// TIA Portal project "EdgeHowTos" (V16) (continued)
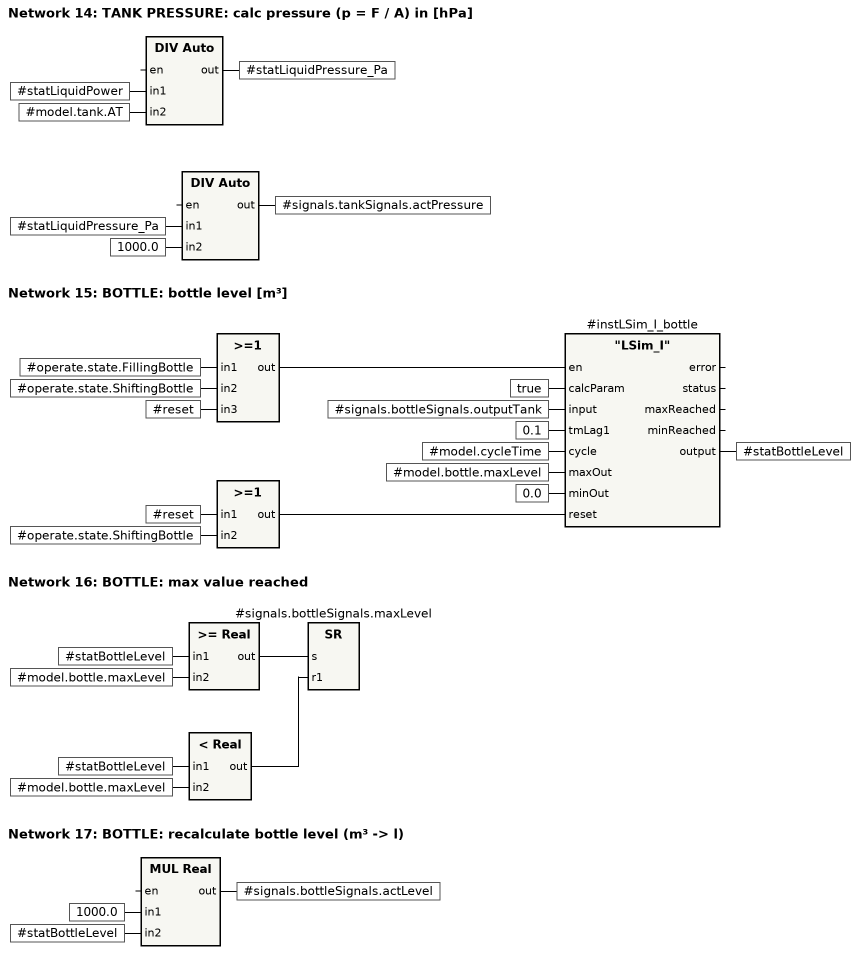
   #statLiquidPressure_Pa := #statLiquidPower / #model.tank.AT;
   #signals.tankSignals.actPressure := #statLiquidPressure_Pa / 1000.0;
END_REGION

REGION Network 15: BOTTLE: bottle level [m³]
   IF #operate.state.FillingBottle OR #operate.state.ShiftingBottle OR #reset THEN
       #instLSim_I_bottle(calcParam := true,   // "LSim_I"
                          input := #signals.bottleSignals.outputTank,
                          tmLag1 := 0.1,
                          cycle := #model.cycleTime,
                          maxOut := #model.bottle.maxLevel,
                          minOut := 0.0,
                          reset := #reset OR #operate.state.ShiftingBottle,
                          output => #statBottleLevel);
   END_IF;
END_REGION

REGION Network 16: BOTTLE: max value reached
   IF #statBottleLevel >= #model.bottle.maxLevel THEN
       #signals.bottleSignals.maxLevel := TRUE;   // SR flip-flop
   END_IF;
   IF #statBottleLevel < #model.bottle.maxLevel THEN #signals.bottleSignals.maxLevel := FALSE; END_IF;
END_REGION

REGION Network 17: BOTTLE: recalculate bottle level (m³ -> l)
   #signals.bottleSignals.actLevel := 1000.0 * #statBottleLevel;
END_REGION

REGION Network 18: HEAT: set init values
   // default value (statHeatingActive = false)
   // - temp = 20°C
   // - tmLag = 0.01
   // (set PT1 controller to initial temperature, otherwise PT1 controller would always start at 0°C)
   // 
   // heating phase (statHeatingActive = true)
   // - temp = 80°C
   // - tmLag = 1
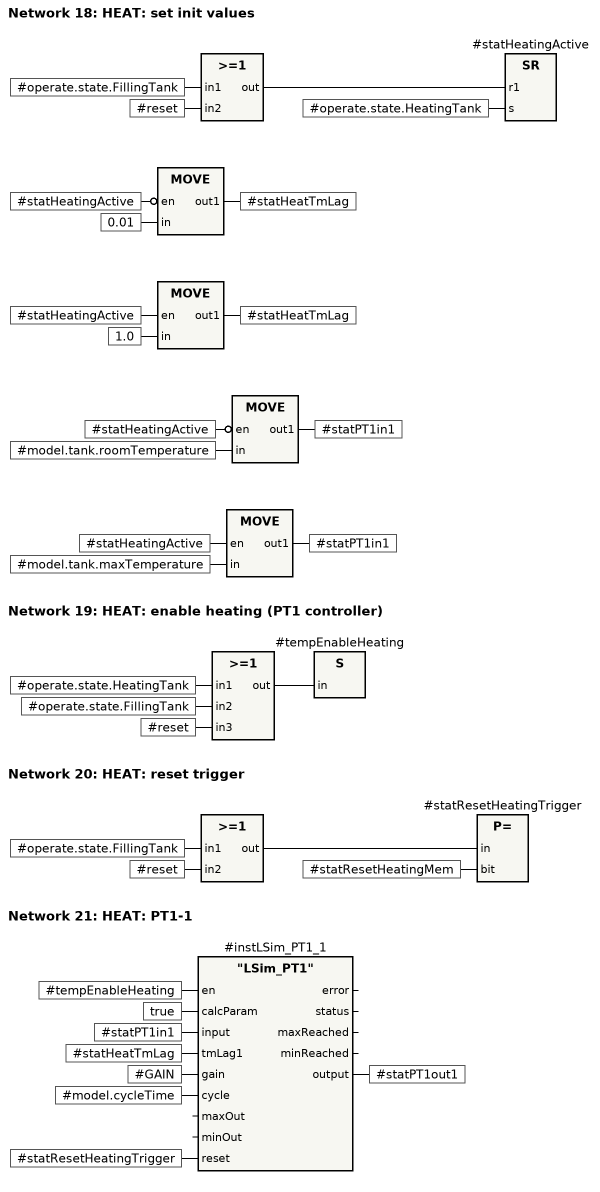
   IF #operate.state.HeatingTank THEN
       #statHeatingActive := TRUE;   // SR flip-flop
   END_IF;
   IF #operate.state.FillingTank OR #reset THEN #statHeatingActive := FALSE; END_IF;
   IF NOT #statHeatingActive THEN #statHeatTmLag := 0.01; END_IF;
   IF #statHeatingActive THEN #statHeatTmLag := 1.0; END_IF;
   IF NOT #statHeatingActive THEN #statPT1in1 := #model.tank.roomTemperature; END_IF;
   IF #statHeatingActive THEN #statPT1in1 := #model.tank.maxTemperature; END_IF;
END_REGION

REGION Network 19: HEAT: enable heating (PT1 controller)
   IF #operate.state.HeatingTank OR #operate.state.FillingTank OR #reset THEN
       #tempEnableHeating := TRUE;
   END_IF;
END_REGION

REGION Network 20: HEAT: reset trigger
   #_w1 := #operate.state.FillingTank OR #reset;
   #statResetHeatingTrigger := #_w1 AND NOT #statResetHeatingMem;   // rising edge
   #statResetHeatingMem := #_w1;
END_REGION

REGION Network 21: HEAT: PT1-1
   IF #tempEnableHeating THEN
       #instLSim_PT1_1(calcParam := true,   // "LSim_PT1"
                       input := #statPT1in1,
                       tmLag1 := #statHeatTmLag,
                       gain := #GAIN,
                       cycle := #model.cycleTime,
                       reset := #statResetHeatingTrigger,
                       output => #statPT1out1);
   END_IF;
END_REGION

REGION Network 22: HEAT: PT1-2
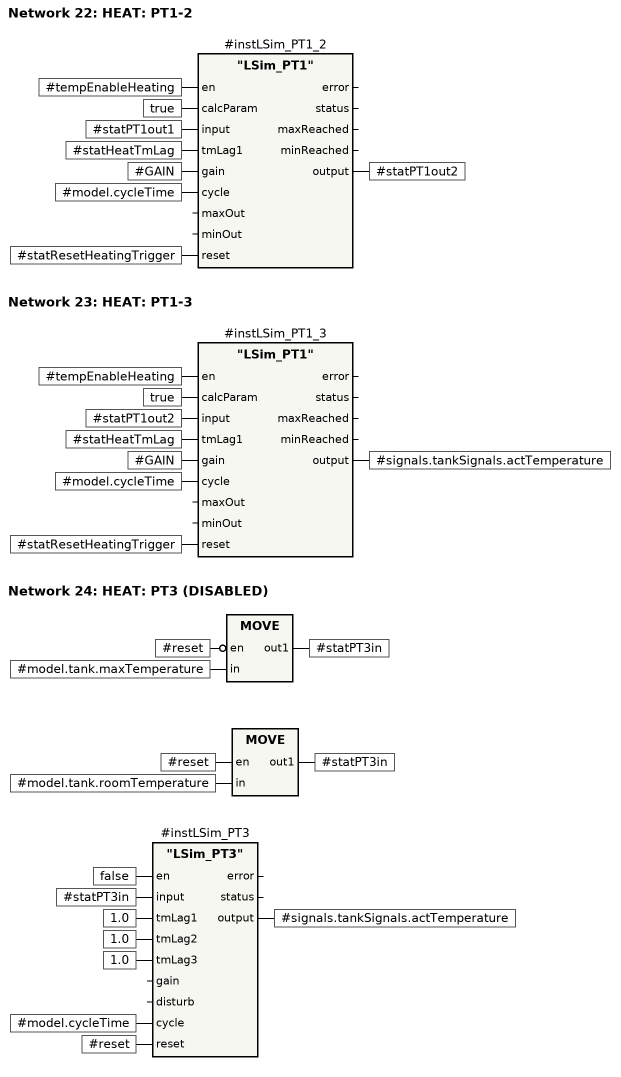
   IF #tempEnableHeating THEN
       #instLSim_PT1_2(calcParam := true,   // "LSim_PT1"
                       input := #statPT1out1,
                       tmLag1 := #statHeatTmLag,
                       gain := #GAIN,
                       cycle := #model.cycleTime,
                       reset := #statResetHeatingTrigger,
                       output => #statPT1out2);
   END_IF;
END_REGION

REGION Network 23: HEAT: PT1-3
   IF #tempEnableHeating THEN
       #instLSim_PT1_3(calcParam := true,   // "LSim_PT1"
                       input := #statPT1out2,
                       tmLag1 := #statHeatTmLag,
                       gain := #GAIN,
                       cycle := #model.cycleTime,
                       reset := #statResetHeatingTrigger,
                       output => #signals.tankSignals.actTemperature);
   END_IF;
END_REGION

REGION Network 24: HEAT: PT3 (DISABLED)
   IF NOT #reset THEN #statPT3in := #model.tank.maxTemperature; END_IF;
   IF #reset THEN #statPT3in := #model.tank.roomTemperature; END_IF;
   IF false THEN
       #instLSim_PT3(input := #statPT3in,   // "LSim_PT3"
                     tmLag1 := 1.0,
                     tmLag2 := 1.0,
                     tmLag3 := 1.0,
                     cycle := #model.cycleTime,
                     reset := #reset,
                     output => #signals.tankSignals.actTemperature);
   END_IF;
END_REGION

REGION Network 25: HEAT: max value reached
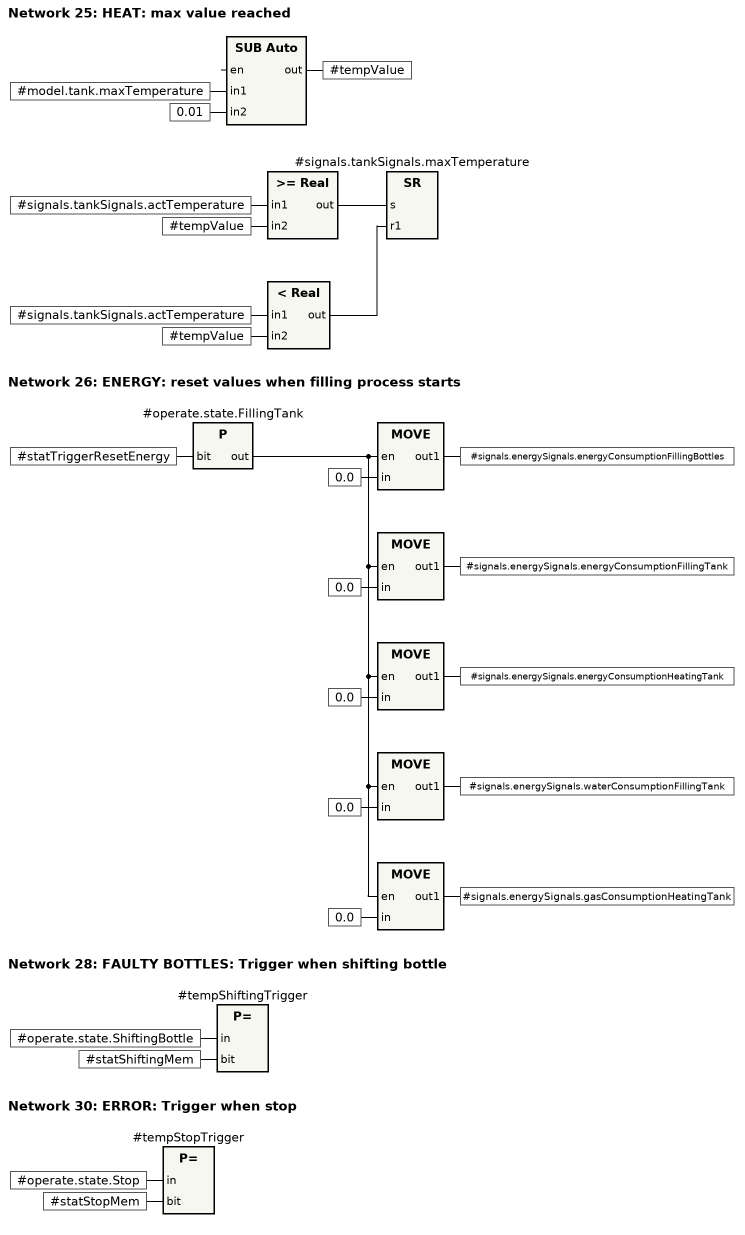
   #tempValue := #model.tank.maxTemperature - 0.01;
   IF #signals.tankSignals.actTemperature >= #tempValue THEN
       #signals.tankSignals.maxTemperature := TRUE;   // SR flip-flop
   END_IF;
   IF #signals.tankSignals.actTemperature < #tempValue THEN
       #signals.tankSignals.maxTemperature := FALSE;
   END_IF;
END_REGION

REGION Network 26: ENERGY: reset values when filling process starts
   #_w1 := #operate.state.FillingTank AND NOT #statTriggerResetEnergy;   // rising edge of #operate.state.FillingTank
   #statTriggerResetEnergy := #operate.state.FillingTank;
   IF #_w1 THEN
       #signals.energySignals.energyConsumptionFillingBottles := 0.0;
       #signals.energySignals.energyConsumptionFillingTank := 0.0;
       #signals.energySignals.energyConsumptionHeatingTank := 0.0;
       #signals.energySignals.waterConsumptionFillingTank := 0.0;
       #signals.energySignals.gasConsumptionHeatingTank := 0.0;
   END_IF;
END_REGION

REGION Network 27 (SCL): ENERGY: calculate values
   // generate random values for energy / water / gas consumption
   // energy [Wh] and water [l] consumption during filling tank
   // ----------------------------------------------------------
   IF #operate.state.FillingTank THEN
       "Random_Number"(Min := 10,
                       Max := 20,
                       RandomNumber => #tempRandomNumber);
       #tempRandomNumber := #tempRandomNumber / 100;
       #signals.energySignals.energyConsumptionFillingTank := #signals.energySignals.energyConsumptionFillingTank + #tempRandomNumber;
       #signals.energySignals.waterConsumptionFillingTank := #signals.tankSignals.actLevel;
   END_IF;

   // energy and gas consumption during heating tank [Wh]
   // ---------------------------------------------------
   IF #operate.state.HeatingTank THEN
       "Random_Number"(Min := 1,
                       Max := 8,
                       RandomNumber => #tempRandomNumber1);
       #tempRandomNumber1 := #tempRandomNumber1 / 10;
       #signals.energySignals.energyConsumptionHeatingTank := #signals.energySignals.energyConsumptionHeatingTank + #tempRandomNumber1;
       #signals.energySignals.gasConsumptionHeatingTank := #signals.energySignals.gasConsumptionHeatingTank + (#tempRandomNumber1 * 1.5);
   END_IF;

   // energy consumption during filling bottles [Wh]
   // -----------------------------------------------
   IF #operate.state.FillingBottle OR #operate.state.ShiftingBottle THEN
       "Random_Number"(Min := 10,
                       Max := 50,
                       RandomNumber => #tempRandomNumber2);
       #tempRandomNumber2 := #tempRandomNumber2 / 100;
       #signals.energySignals.energyConsumptionFillingBottles := #signals.energySignals.energyConsumptionFillingBottles + #tempRandomNumber2;
   END_IF;
END_REGION

REGION Network 28: FAULTY BOTTLES: Trigger when shifting bottle
   #tempShiftingTrigger := #operate.state.ShiftingBottle AND NOT #statShiftingMem;   // rising edge
   #statShiftingMem := #operate.state.ShiftingBottle;
END_REGION

REGION Network 29 (SCL): FAULTY BOTTLES: Simulate faulty bottles (generate random number)
   IF #tempShiftingTrigger THEN
       "Random_Number"(Min := 0,
                       Max := 8,
                       RandomNumber => #tempRandomNumber3);

       IF (#tempRandomNumber3 = 1) OR (#tempRandomNumber3 = 5) THEN
           #process.numberFaulty := #process.numberFaulty + 1;
       END_IF;

   END_IF;
END_REGION

REGION Network 30: ERROR: Trigger when stop
   #tempStopTrigger := #operate.state.Stop AND NOT #statStopMem;   // rising edge
   #statStopMem := #operate.state.Stop;
END_REGION

REGION Network 31 (SCL): ERROR: Simulate error
       IF #errors.errorSimulation THEN

           // random error generation
           IF #tempShiftingTrigger THEN
               "Random_Number"(Min := 0,
                               Max := 100,
                               RandomNumber => #tempRandomNumber5);

               // go into error state
               IF #tempRandomNumber5 = 1 THEN
                   #appSignals.APP_Error := true;
               END_IF;

           END_IF;

           // triggered error genertion
           IF #errors.errorTrigger THEN
               #appSignals.APP_Error := true;
           END_IF;


           // if timer finished (negative edge on it's output), go in stop > start again
           "F_TRIG_DB_Error_Finished"(CLK := #instTimerError.Q,
                                      Q => #statResetError);

           // reset error > machine goes automatically into stop
           IF #statResetError THEN
               #appSignals.APP_Error := false;
               #errors.errorCode := "ERROR_0_NO";
               #statResetError := false;
               #statStart := true;
           END_IF;

           IF #tempStopTrigger AND #statStart THEN
               #appSignals.APP_Start := true;
               #statStart := false;
           END_IF;

       END_IF;
END_REGION

REGION Network 32: ERROR: Trigger when new error comes in and start timer
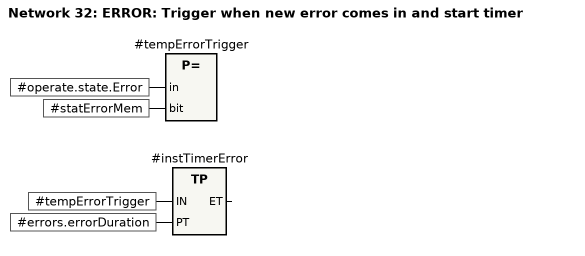
   #tempErrorTrigger := #operate.state.Error AND NOT #statErrorMem;   // rising edge
   #statErrorMem := #operate.state.Error;
   #instTimerError.TP(IN := #tempErrorTrigger, PT := #errors.errorDuration);
END_REGION

REGION Network 33 (SCL): ERROR: Simulate error codes
   // Codes btw. 1-6 (7 = HMI error)
   IF #errors.errorSimulation THEN

       // generate random error code
       IF #tempErrorTrigger AND (#errors.errorCode = "ERROR_0_NO") THEN

           "Random_Number"(Min := 1,
                           Max := 6,
                           RandomNumber => #tempRandomNumber4);

           #errors.errorCode := #tempRandomNumber4;

       END_IF;

   END_IF;
END_REGION
END_FUNCTION_BLOCK

FUNCTION_BLOCK "LSim_PT1"   // FB50, SCL
{ S7_Optimized_Access := 'TRUE' }
VERSION : 2.01
   VAR_INPUT
      calcParam : Bool;   // recalculate with new parameters
      input : Real;   // input signal
      tmLag1 : Real := 1.0;   // time constant T1 [sec]
      gain : Real := 1.0;   // gain factor
      cycle : Real := 0.1;   // cyclic time [sec]
      maxOut : Real := 100.0;   // max. output limit
      minOut : Real;   // min. output limit
      reset : Bool;   // resets all relevant parameters to ‘0’ including the output
   END_VAR
   VAR_OUTPUT
      error : Bool;   // error (#tmLag1 <= 0)
      status : Word;   // status (if #tmLag1 <= 0 then status = 16#8001)
      maxReached : Bool;   // output has reached max. limit
      minReached : Bool;   // output has reached min. limit
      output : Real;   // output signal (if #error = FALSE)
   END_VAR
   VAR
      statRf1 : Real;
      statRe1 : Real;
      statOverfirst : Bool;
      statOutput : Real;
   END_VAR
BEGIN
   //=============================================================================
   //SIEMENS AG
   //(c)Copyright 2017 All Rights Reserved
   //-----------------------------------------------------------------------------
   //Library:       Library for Controlled System Simulation
   //Tested with:   S7-1500 FW V2.0 / S7-1200 FW V4.2
   //Engineering:   STEP 7 V14 Upd2 (TIA Portal)
   //Restrictions:  Cyclic interrupt
   //Requirements:  memory card needed for S7-1500
   //Functionality: Simulation of a PT1-System
   //
   //              gain
   //  F(p) = ---------------
   //          tmLag1 * p + 1
   //          
   //  Call the simulation in a cyclic interrupt with
   //  cyclic interrupt time at least = tmLag1/10!
   //-----------------------------------------------------------------------------
   //Change log table:
   //Version  Date       Expert in charge                Changes applied
   //02.00.00 03.02.2016 Siemens Industry Online Support Release (STEP 7 V13 SP1)
   //02.00.01 02.03.2017 Siemens Industry Online Support Release (STEP 7 V14)
   //=============================================================================
   // check parameter
   IF #tmLag1 <= 0 THEN
     #error := TRUE;
     #status := W#16#8001;     // Parameter Error
     #statOutput := 0;
     #output := 0;
     RETURN;
   ELSE
     #error := FALSE;
     #status := W#16#0000;     // no error
   END_IF;

   IF #calcParam = True OR NOT #statOverfirst THEN
     #statOverfirst:=1;
   // Z-parameters For Laplace PT1-System
   #statRe1 := - EXP(-#cycle/#tmLag1);
   #statRf1 := #gain*(1 + #statRe1);
   END_IF;

   // Differencial Equation of PT1-System
   #statOutput := #input*#statRf1 - #statOutput*#statRe1;

   // max limit of acutating variable
   IF #statOutput > #maxOut THEN
     #statOutput := #maxOut;
     #maxReached:= True;
   ELSE
     #maxReached := False;
   END_IF;

   // min limit of acutating variable
   IF #statOutput < #minOut THEN
     #statOutput := #minOut;
     #minReached := True;
   ELSE
     #minReached := False;
   END_IF;

   IF #reset THEN
     #statOutput := 0;
   END_IF;

   #output := #statOutput;
END_FUNCTION_BLOCK

FUNCTION_BLOCK "LSim_PT3"   // FB54, SCL
{ S7_Optimized_Access := 'TRUE' }
VERSION : 2.01
   VAR_INPUT
      input : Real;   // input variable
      tmLag1 : Real := 29.0;   // time lag 1 in s
      tmLag2 : Real := 17.5;   // time lag 2 in s
      tmLag3 : Real := 3.1;   // time lag 3 in s
      gain : Real := 1.0;   // proportional gain
      disturb : Real;   // disturbance variable (additional to "input")
      cycle : Real := 0.1;   // sample time [in sec]
      reset : Bool;   // complete restart (#output = #input)
   END_VAR
   VAR_OUTPUT
      error : Bool;   // error (#tmLag1 <= 0 or #tmLag2 <= 0 or #tmLag3 <= 0)
      status : Word;   // status (if #error = TRUE then status = 16#8001)
      output : Real;   // output signal (if #error = FALSE)
   END_VAR
   VAR
      statFback1 : Real;   // feedback path value 1
      statFback2 : Real;   // feedback path value 2
      statFback3 : Real;   // feedback path value 3
   END_VAR
   VAR_TEMP
      tempHvar : Real;   // help variable
      tempCycleR : Real;   // cycle to real
      tempTmLag1R : Real;   // time lag 1 to real
      tempTmLag2R : Real;   // time lag 2 to real
      tempTmLag3R : Real;   // time lag 3 to real
      tempOutvNew : Real;   // new output variable
   END_VAR
BEGIN
   //=============================================================================
   //SIEMENS AG
   //(c)Copyright 2017 All Rights Reserved
   //-----------------------------------------------------------------------------
   //Library:       Library for Controlled System Simulation
   //Tested with:   S7-1500 FW V2.0 / S7-1200 FW V4.2
   //Engineering:   STEP 7 V14 Upd2 (TIA Portal)
   //Restrictions:  Cyclic interrupt
   //Requirements:  memory card needed for S7-1500
   //Functionality: Simulation of an PT3-system
   //
   //                               gain
   //  F(p) = ------------------------------------------------------
   //         (tmLag1 * p + 1) * (tmLag2 * p + 1) * (tmLag3 * p + 1)
   //          
   //  Call the simulation in a cyclic interrupt with
   //  cyclic interrupt time at least = tmLag1/10!
   //-----------------------------------------------------------------------------
   //Change log table:
   //Version  Date       Expert in charge                Changes applied
   //02.00.00 03.02.2016 Siemens Industry Online Support Release (STEP 7 V13 SP1)
   //02.00.01 02.03.2017 Siemens Industry Online Support Release (STEP 7 V14)
   //=============================================================================
   // check parameter
   IF #tmLag1 <= 0 OR #tmLag2 <= 0 OR #tmLag3 <= 0 THEN
     #error := TRUE;
     #status := W#16#8001;     // Parameter Error
     #output := #input; //write output data
     #statFback1 := #input; //write static data
     #statFback2 := #input;
     #statFback3 := #input;
     RETURN;
   ELSE
     #error := FALSE;
     #status := W#16#0000;     // no error
   END_IF;

   IF #reset THEN //complete restart routine

     #output := #input;//write output data
     #statFback1 := #input;//write static data
     #statFback2 := #input;
     #statFback3 := #input;

   ELSE //cycle mode routine

     #tempCycleR  := #cycle*1000; //transform data type
     #tempTmLag1R := #tmLag1*1000;
     #tempTmLag2R := #tmLag2*1000;
     #tempTmLag3R := #tmLag3*1000;

     IF #tempCycleR * 0.5 > #tempTmLag1R THEN //limit TM_LAG1
       #tempTmLag1R := #tempCycleR * 0.5;
     END_IF;

     IF #tempCycleR * 0.5 > #tempTmLag2R THEN //limit TM_LAG2
       #tempTmLag2R := #tempCycleR * 0.5;
     END_IF;

     IF #tempCycleR * 0.5 > #tempTmLag3R THEN //limit TM_LAG2
       #tempTmLag3R := #tempCycleR * 0.5;
     END_IF;

     //1. first order lag algorithm
     #tempHvar     := #tempCycleR / (#tempTmLag1R * 2.0); 
     #tempHvar     := (#gain * (#input + #disturb) - #statFback1) * #tempHvar / (#tempHvar + 1.0);
     #tempOutvNew  := #tempHvar + #statFback1;
     #statFback1  := #tempHvar * 2.0 + #statFback1;

     //2. first order lag algorithm
     #tempHvar     := #tempCycleR / (#tempTmLag2R * 2.0); 
     #tempHvar     := ((#tempOutvNew - #statFback2) * #tempHvar) / (#tempHvar + 1.0);
     #tempOutvNew  := #tempHvar + #statFback2;
     #statFback2  := #tempHvar * 2.0 + #statFback2;

     //3. first order lag algorithm
     #tempHvar     := #tempCycleR / (#tempTmLag3R * 2.0); 
     #tempHvar     := ((#tempOutvNew - #statFback3) * #tempHvar) / (#tempHvar + 1.0);
     #tempOutvNew  := #tempHvar + #statFback3;
     #statFback3  := #tempHvar * 2.0 + #statFback3;

     #output := #tempOutvNew; //write output

   END_IF;
END_FUNCTION_BLOCK

FUNCTION_BLOCK "LSim_I"   // FB56, SCL
{ S7_Optimized_Access := 'TRUE' }
VERSION : 2.01
   VAR_INPUT
      calcParam : Bool;   // recalculate with new parameters
      input : Real;   // input signal
      tmLag1 : Real := 1.0;   // time constant T1 [sec]
      cycle : Real := 0.1;   // cyclic time [sec]
      maxOut : Real := 100.0;   // max. output limit
      minOut : Real;   // min. output limit
      reset : Bool;   // resets all relevant parameters to ‘0’ including the output
   END_VAR
   VAR_OUTPUT
      error : Bool;   // error (#tmLag1 <= 0)
      status : Word;   // status (if #tmLag1 <= 0 then status = 16#8001)
      maxReached : Bool;   // output has reached max. limit
      minReached : Bool;   // output has reached min. limit
      output : Real;   // output signal (if #error = FALSE)
   END_VAR
   VAR
      statRxn1 : Real;   // delayed input signal (n-1)
      statRyn1 : Real;   // delayed output signal (n-1)
      statRa1 : Real;
      statRb1 : Real;
      statOverfirst : Bool;
      statOutput : Real;   // output signal
   END_VAR
BEGIN
   //=============================================================================
   //SIEMENS AG
   //(c)Copyright 2017 All Rights Reserved
   //-----------------------------------------------------------------------------
   //Library:       Library for Controlled System Simulation
   //Tested with:   S7-1500 FW V2.0 / S7-1200 FW V4.2
   //Engineering:   STEP 7 V14 Upd2 (TIA Portal)
   //Restrictions:  Cyclic interrupt
   //Requirements:  memory card needed for S7-1500
   //Functionality: Simulation of a I-System
   //
   //             1
   //  F(p) = -----------
   //         (tmLag1*p)
   //          
   //  Call the simulation in a cyclic interrupt with
   //  cyclic interrupt time at least = tmLag1/10!
   //-----------------------------------------------------------------------------
   //Change log table:
   //Version  Date       Expert in charge                Changes applied
   //02.00.00 03.02.2016 Siemens Industry Online Support Release (STEP 7 V13 SP1)
   //02.00.01 02.03.2017 Siemens Industry Online Support Release (STEP 7 V14)
   //=============================================================================

   // check parameter
   IF #tmLag1 <= 0 THEN
     #error := True;
     #status := W#16#8001;     // Parameter Error
     #statRxn1 := 0.0;
     #statRyn1 := 0.0;
     #statOutput := 0;
     #output := 0;
     RETURN;
   ELSE
     #error := FALSE;
     #status := W#16#0000;     // no error
   END_IF;

   // calculates the z-parameter for the difference equatation
   IF #calcParam = True OR NOT #statOverfirst THEN
   #statOverfirst:=1;
     // Calculate z-parameters for IT1-System
   #statRb1 := #cycle/#tmLag1;
   #statRa1 := -1;

   END_IF;

   // reset Memory
   IF #reset = True THEN
     #statRxn1 := 0.0;
     #statRyn1 := 0.0;
     #statOutput:=0;
   END_IF;

   // save delayed output-signals
   #statRyn1:= #statOutput;

   // difference equatation for the I-system
   #statOutput := #statRxn1* #statRb1 - #statRyn1*#statRa1;

   // save delayed input-signals
   #statRxn1 := #input;

   // max limit of acutating variable
   IF #statOutput > #maxOut THEN
     #statOutput := #maxOut;
     #maxReached:= True;
   ELSE
     #maxReached := False;
   END_IF;